REGION Network 19: QW98 - Spare Output (Hardware Channel De-activated)
   RUNG wire#powerrail
      P_Contact(operand := "80_From_HMI".MAN_AQ_INC_98, bit := "90_Manual_Data".INC_PLS_98)
      wire#w1
      Add(in1 := "16_AQ_Data".R2_SPR_AQ_98, in2 := 1.0, out => "16_AQ_Data".R2_SPR_AQ_98)
      { S7_Templates := "SrcType := Real" } GE_Contact(in1 := "16_AQ_Data".R2_SPR_AQ_98, in2 := "16_AQ_Data".QW_98.ENG_MAX)
      { S7_GenerateENO := "TRUE" } Move(in := "16_AQ_Data".QW_98.ENG_MAX, out1 => "16_AQ_Data".R2_SPR_AQ_98)
   END_RUNG
   RUNG wire#powerrail
      Contact( "80_From_HMI".MAN_AQ_INC_98 )
      P_Contact(operand := "Clock_5Hz", bit := "90_Manual_Data".INC_PLS_98_Hz)
   END_RUNG wire#w1
   RUNG wire#powerrail
      P_Contact(operand := "80_From_HMI".MAN_AQ_DEC_98, bit := "90_Manual_Data".DEC_PLS_98)
      wire#w2
      Sub(in1 := "16_AQ_Data".R2_SPR_AQ_98, in2 := 1.0, out => "16_AQ_Data".R2_SPR_AQ_98)
      { S7_Templates := "SrcType := Real" } LE_Contact(in1 := "16_AQ_Data".R2_SPR_AQ_98, in2 := "16_AQ_Data".QW_98.ENG_MIN)
      { S7_GenerateENO := "TRUE" } Move(in := "16_AQ_Data".QW_98.ENG_MIN, out1 => "16_AQ_Data".R2_SPR_AQ_98)
   END_RUNG
   RUNG wire#powerrail
      Contact( "80_From_HMI".MAN_AQ_DEC_98 )
      P_Contact(operand := "Clock_5Hz", bit := "90_Manual_Data".DEC_PLS_98_Hz)
   END_RUNG wire#w2
   // the same network as SCL:
   #_w1 := "80_From_HMI".MAN_AQ_INC_98 AND NOT "90_Manual_Data".INC_PLS_98;   // rising edge of "80_From_HMI".MAN_AQ_INC_98
   "90_Manual_Data".INC_PLS_98 := "80_From_HMI".MAN_AQ_INC_98;
   #_w2 := "80_From_HMI".MAN_AQ_INC_98 AND "Clock_5Hz" AND NOT "90_Manual_Data".INC_PLS_98_Hz;   // rising edge of "Clock_5Hz"
   "90_Manual_Data".INC_PLS_98_Hz := "Clock_5Hz";
   #_w3 := #_w1 OR #_w2;
   IF #_w3 THEN "16_AQ_Data".R2_SPR_AQ_98 := "16_AQ_Data".R2_SPR_AQ_98 + 1.0; END_IF;
   IF #_w3 AND ("16_AQ_Data".R2_SPR_AQ_98 >= "16_AQ_Data".QW_98.ENG_MAX) THEN
       "16_AQ_Data".R2_SPR_AQ_98 := "16_AQ_Data".QW_98.ENG_MAX;
   END_IF;
   #_w4 := "80_From_HMI".MAN_AQ_DEC_98 AND NOT "90_Manual_Data".DEC_PLS_98;   // rising edge of "80_From_HMI".MAN_AQ_DEC_98
   "90_Manual_Data".DEC_PLS_98 := "80_From_HMI".MAN_AQ_DEC_98;
   #_w5 := "80_From_HMI".MAN_AQ_DEC_98 AND "Clock_5Hz" AND NOT "90_Manual_Data".DEC_PLS_98_Hz;   // rising edge of "Clock_5Hz"
   "90_Manual_Data".DEC_PLS_98_Hz := "Clock_5Hz";
   #_w6 := #_w4 OR #_w5;
   IF #_w6 THEN "16_AQ_Data".R2_SPR_AQ_98 := "16_AQ_Data".R2_SPR_AQ_98 - 1.0; END_IF;
   IF #_w6 AND ("16_AQ_Data".R2_SPR_AQ_98 <= "16_AQ_Data".QW_98.ENG_MIN) THEN
       "16_AQ_Data".R2_SPR_AQ_98 := "16_AQ_Data".QW_98.ENG_MIN;
   END_IF;
END_REGION

REGION Network 20: QW100 - Main Fuel Reg Valve Control (CV-203)
   RUNG wire#powerrail
      P_Contact(operand := "80_From_HMI".MAN_AQ_INC_100, bit := "90_Manual_Data".INC_PLS_100)
      wire#w1
      Add(in1 := "16_AQ_Data".CV203_CNTRL, in2 := 1.0, out => "16_AQ_Data".CV203_CNTRL)
      { S7_Templates := "SrcType := Real" } GE_Contact(in1 := "16_AQ_Data".CV203_CNTRL, in2 := "16_AQ_Data".QW_100.ENG_MAX)
      { S7_GenerateENO := "TRUE" } Move(in := "16_AQ_Data".QW_100.ENG_MAX, out1 => "16_AQ_Data".CV203_CNTRL)
   END_RUNG
   RUNG wire#powerrail
      Contact( "80_From_HMI".MAN_AQ_INC_100 )
      P_Contact(operand := "Clock_5Hz", bit := "90_Manual_Data".INC_PLS_100_Hz)
   END_RUNG wire#w1
   RUNG wire#powerrail
      P_Contact(operand := "80_From_HMI".MAN_AQ_DEC_100, bit := "90_Manual_Data".DEC_PLS_100)
      wire#w2
      Sub(in1 := "16_AQ_Data".CV203_CNTRL, in2 := 1.0, out => "16_AQ_Data".CV203_CNTRL)
      { S7_Templates := "SrcType := Real" } LE_Contact(in1 := "16_AQ_Data".CV203_CNTRL, in2 := "16_AQ_Data".QW_100.ENG_MIN)
      { S7_GenerateENO := "TRUE" } Move(in := "16_AQ_Data".QW_100.ENG_MIN, out1 => "16_AQ_Data".CV203_CNTRL)
   END_RUNG
   RUNG wire#powerrail
      Contact( "80_From_HMI".MAN_AQ_DEC_100 )
      P_Contact(operand := "Clock_5Hz", bit := "90_Manual_Data".DEC_PLS_100_Hz)
   END_RUNG wire#w2
   // the same network as SCL:
   #_w1 := "80_From_HMI".MAN_AQ_INC_100 AND NOT "90_Manual_Data".INC_PLS_100;   // rising edge of "80_From_HMI".MAN_AQ_INC_100
   "90_Manual_Data".INC_PLS_100 := "80_From_HMI".MAN_AQ_INC_100;
   #_w2 := "80_From_HMI".MAN_AQ_INC_100 AND "Clock_5Hz" AND NOT "90_Manual_Data".INC_PLS_100_Hz;   // rising edge of "Clock_5Hz"
   "90_Manual_Data".INC_PLS_100_Hz := "Clock_5Hz";
   #_w3 := #_w1 OR #_w2;
   IF #_w3 THEN "16_AQ_Data".CV203_CNTRL := "16_AQ_Data".CV203_CNTRL + 1.0; END_IF;
   IF #_w3 AND ("16_AQ_Data".CV203_CNTRL >= "16_AQ_Data".QW_100.ENG_MAX) THEN
       "16_AQ_Data".CV203_CNTRL := "16_AQ_Data".QW_100.ENG_MAX;
   END_IF;
   #_w4 := "80_From_HMI".MAN_AQ_DEC_100 AND NOT "90_Manual_Data".DEC_PLS_100;   // rising edge of "80_From_HMI".MAN_AQ_DEC_100
   "90_Manual_Data".DEC_PLS_100 := "80_From_HMI".MAN_AQ_DEC_100;
   #_w5 := "80_From_HMI".MAN_AQ_DEC_100 AND "Clock_5Hz" AND NOT "90_Manual_Data".DEC_PLS_100_Hz;   // rising edge of "Clock_5Hz"
   "90_Manual_Data".DEC_PLS_100_Hz := "Clock_5Hz";
   #_w6 := #_w4 OR #_w5;
   IF #_w6 THEN "16_AQ_Data".CV203_CNTRL := "16_AQ_Data".CV203_CNTRL - 1.0; END_IF;
   IF #_w6 AND ("16_AQ_Data".CV203_CNTRL <= "16_AQ_Data".QW_100.ENG_MIN) THEN
       "16_AQ_Data".CV203_CNTRL := "16_AQ_Data".QW_100.ENG_MIN;
   END_IF;
END_REGION

REGION Network 21: QW102 - Main Atom Air Reg Valve Control (CV-111)
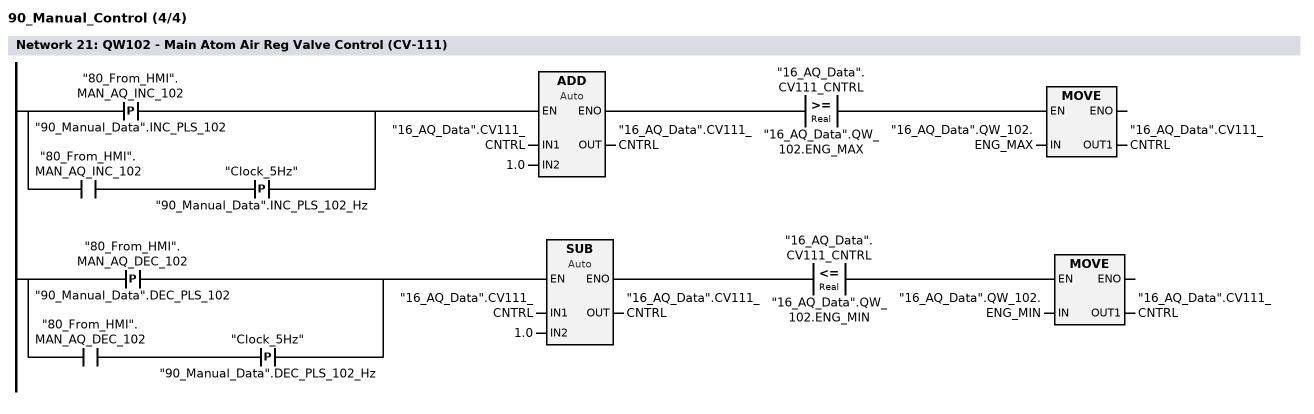
   RUNG wire#powerrail
      P_Contact(operand := "80_From_HMI".MAN_AQ_INC_102, bit := "90_Manual_Data".INC_PLS_102)
      wire#w1
      Add(in1 := "16_AQ_Data".CV111_CNTRL, in2 := 1.0, out => "16_AQ_Data".CV111_CNTRL)
      { S7_Templates := "SrcType := Real" } GE_Contact(in1 := "16_AQ_Data".CV111_CNTRL, in2 := "16_AQ_Data".QW_102.ENG_MAX)
      { S7_GenerateENO := "TRUE" } Move(in := "16_AQ_Data".QW_102.ENG_MAX, out1 => "16_AQ_Data".CV111_CNTRL)
   END_RUNG
   RUNG wire#powerrail
      Contact( "80_From_HMI".MAN_AQ_INC_102 )
      P_Contact(operand := "Clock_5Hz", bit := "90_Manual_Data".INC_PLS_102_Hz)
   END_RUNG wire#w1
   RUNG wire#powerrail
      P_Contact(operand := "80_From_HMI".MAN_AQ_DEC_102, bit := "90_Manual_Data".DEC_PLS_102)
      wire#w2
      Sub(in1 := "16_AQ_Data".CV111_CNTRL, in2 := 1.0, out => "16_AQ_Data".CV111_CNTRL)
      { S7_Templates := "SrcType := Real" } LE_Contact(in1 := "16_AQ_Data".CV111_CNTRL, in2 := "16_AQ_Data".QW_102.ENG_MIN)
      { S7_GenerateENO := "TRUE" } Move(in := "16_AQ_Data".QW_102.ENG_MIN, out1 => "16_AQ_Data".CV111_CNTRL)
   END_RUNG
   RUNG wire#powerrail
      Contact( "80_From_HMI".MAN_AQ_DEC_102 )
      P_Contact(operand := "Clock_5Hz", bit := "90_Manual_Data".DEC_PLS_102_Hz)
   END_RUNG wire#w2
   // the same network as SCL:
   #_w1 := "80_From_HMI".MAN_AQ_INC_102 AND NOT "90_Manual_Data".INC_PLS_102;   // rising edge of "80_From_HMI".MAN_AQ_INC_102
   "90_Manual_Data".INC_PLS_102 := "80_From_HMI".MAN_AQ_INC_102;
   #_w2 := "80_From_HMI".MAN_AQ_INC_102 AND "Clock_5Hz" AND NOT "90_Manual_Data".INC_PLS_102_Hz;   // rising edge of "Clock_5Hz"
   "90_Manual_Data".INC_PLS_102_Hz := "Clock_5Hz";
   #_w3 := #_w1 OR #_w2;
   IF #_w3 THEN "16_AQ_Data".CV111_CNTRL := "16_AQ_Data".CV111_CNTRL + 1.0; END_IF;
   IF #_w3 AND ("16_AQ_Data".CV111_CNTRL >= "16_AQ_Data".QW_102.ENG_MAX) THEN
       "16_AQ_Data".CV111_CNTRL := "16_AQ_Data".QW_102.ENG_MAX;
   END_IF;
   #_w4 := "80_From_HMI".MAN_AQ_DEC_102 AND NOT "90_Manual_Data".DEC_PLS_102;   // rising edge of "80_From_HMI".MAN_AQ_DEC_102
   "90_Manual_Data".DEC_PLS_102 := "80_From_HMI".MAN_AQ_DEC_102;
   #_w5 := "80_From_HMI".MAN_AQ_DEC_102 AND "Clock_5Hz" AND NOT "90_Manual_Data".DEC_PLS_102_Hz;   // rising edge of "Clock_5Hz"
   "90_Manual_Data".DEC_PLS_102_Hz := "Clock_5Hz";
   #_w6 := #_w4 OR #_w5;
   IF #_w6 THEN "16_AQ_Data".CV111_CNTRL := "16_AQ_Data".CV111_CNTRL - 1.0; END_IF;
   IF #_w6 AND ("16_AQ_Data".CV111_CNTRL <= "16_AQ_Data".QW_102.ENG_MIN) THEN
       "16_AQ_Data".CV111_CNTRL := "16_AQ_Data".QW_102.ENG_MIN;
   END_IF;
END_REGION
END_FUNCTION

// ===== PLC "Rack 3 - GCU & BWT PLC - 7KF2"  CPU 1516F-3 PN/DP =====

VAR_GLOBAL   // PLC tag table "Default tag table"
   "Clock_10Hz" AT %M0.0 : Bool;   // System bit
   "Clock_5Hz" AT %M0.1 : Bool;   // System bit
   "Clock_2.5Hz" AT %M0.2 : Bool;   // System bit
   "Clock_2Hz" AT %M0.3 : Bool;   // System bit
   "Clock_1.25Hz" AT %M0.4 : Bool;   // System bit
   "Clock_1Hz" AT %M0.5 : Bool;   // System bit
   "Clock_0.625Hz" AT %M0.6 : Bool;   // System bit
   "Clock_0.5Hz" AT %M0.7 : Bool;   // System bit
   "Clock_Byte" AT %MB0 : Byte;   // System bit
   "System_Byte" AT %MB1 : Byte;   // System bit
   "FirstScan" AT %M1.0 : Bool;   // System bit
   "DiagStatusUpdate" AT %M1.1 : Bool;   // System bit
   "AlwaysTRUE" AT %M1.2 : Bool;   // System bit
   "AlwaysFALSE" AT %M1.3 : Bool;   // System bit
   "Tag_1" AT %M222.2 : Bool;
   "Tag_2" AT %ID222 : Real;
   "Tag_3" AT %ID223 : Real;
   "Tag_4" AT %ID224 : Real;
   "Tag_5" AT %ID221 : Real;
   "Tag_6" AT %M1000.0 : Bool;
   "Tag_7" AT %MD1002 : Real;
   "TEST" AT %M2.0 : Bool;
   "Tag_8" AT %M55.0 : Bool;
   "Tag_9" AT %MD55 : DWord;
   "Tag_10" AT %MD56 : Real;
   "Tag_11" AT %MD57 : Real;
   "Tag_12" AT %MD58 : DWord;
   "Tag_13" AT %MD59 : Real;
   "Tag_14" AT %MD60 : DWord;
   "Tag_15" AT %MD61 : Real;
   "Tag_16" AT %MD62 : DWord;
   "Tag_17" AT %MD63 : Real;
   "Tag_18" AT %MD64 : DWord;
   "Tag_19" AT %MD65 : Real;
   "Tag_20" AT %MD66 : DWord;
   "Tag_21" AT %MD67 : Real;
   "Tag_22" AT %MD68 : DWord;
   "Tag_23" AT %MD69 : DWord;
   "Tag_24" AT %MD70 : Real;
   "Tag_25" AT %MD71 : DWord;
   "Tag_26" AT %MD72 : Real;
   "Tag_27" AT %MD73 : Real;
   "Tag_28" AT %MD74 : DWord;
   "Tag_29" AT %MD75 : Real;
   "Tag_30" AT %MD76 : DWord;
   "Tag_31" AT %MD77 : Real;
   "Tag_32" AT %MD78 : DWord;
   "Tag_33" AT %MD79 : Real;
   "Tag_34" AT %MD80 : DWord;
   "Tag_35" AT %MD81 : Real;
   "Tag_36" AT %MD82 : DWord;
END_VAR

VAR_GLOBAL   // PLC tag table "PLC_IO"
   "R3_SPR_DI_136_0" AT %I136.0 : Bool;   // Spare input
   "R3_SPR_DI_136_1" AT %I136.1 : Bool;   // Spare input
   "Cooling Seawater Flow Switch" AT %I136.2 : Bool;   // FS332-8B1
   "Fresh Water Cooling Flow Switch" AT %I136.5 : Bool;   // FS350-8B3
   "GCU Drain Valve Feedback Open" AT %I136.6 : Bool;   // CV341-8B4
   "GCU Drain Valve Feedback Closed" AT %I136.7 : Bool;   // CV341-8B4
   "Gas to Deck Valve Feedback Open" AT %I137.0 : Bool;   // CV406-9B1
   "Gas to Deck Valve Feedback Closed" AT %I137.1 : Bool;   // CV406-9B1
   "Gas Block Valve 1 Feedback Open" AT %I137.2 : Bool;   // CV407-9B2
   "Gas Block Valve 1 Feedback Closed" AT %I137.3 : Bool;   // CV407-9B2
   "Gas Block Valve 2 Feedback Open" AT %I137.4 : Bool;   // CV411-9B3
   "Gas Block Valve 2 Feedback Closed" AT %I137.5 : Bool;   // CV411-9B3
   "Gas Bleed Valve Feedback Open" AT %I137.6 : Bool;   // CV409-9B4
   "Gas Bleed Valve Feedback Closed" AT %I137.7 : Bool;   // CV409-9B4
   "Ambient Air Valve Feedback Open" AT %I138.0 : Bool;   // CV441-10B1
   "Ambient Air Valve Feedback Closed" AT %I138.1 : Bool;   // CV441-10B1
   "GCU Low Level Switch" AT %I138.2 : Bool;   // LS303-10B2
   "GCU Booster Pump Enabled" AT %I138.3 : Bool;   // P304-MCCP
   "GCU Local PB - Start" AT %I138.4 : Bool;   // 10S1
   "GCU Local PB - Stop" AT %I138.5 : Bool;   // 10S2
   "E-Stop Pressed @ BWT CP" AT %I138.6 : Bool;   // 8S1
   "GCU Recirculation Pump Enabled" AT %I138.7 : Bool;   // P303-MCCP
   "Process Gas Compressor Running/Stopped" AT %I139.0 : Bool;   // E400
   "Process Gas Compressor Tripped/Shutdown" AT %I139.1 : Bool;   // E400
   "GCU Recirculation Pump Healthy" AT %I139.2 : Bool;   // P303-MCCP
   "5T1 Power Healthy" AT %I139.3 : Bool;   // 5T2
   "Panel Vent Power Healthy" AT %I139.4 : Bool;   // 6Q6
   "GCU Booster Pump Healthy" AT %I139.5 : Bool;   // P304-MCCP
   "PGC Running Loaded/On-line" AT %I139.6 : Bool;   // E400
   "PGC Alarm/Warning" AT %I139.7 : Bool;   // E400
   "GCU Level" AT %IW800 : Int;   // LIT304
   "R3_SPR_AI_802" AT %IW802 : Int;   // Spare input
   "Fresh Water Cooling Temperature" AT %IW804 : Int;   // TIT408
   "Gas to Deck (Outlet) Temperature" AT %IW806 : Int;   // TIT406
   "Gas To Deck Vent Valve Feedback" AT %IW808 : Int;   // CV405
   "Gas to Deck Pressure" AT %IW810 : Int;   // PIT416
   "Fresh Water Inlet Pressure" AT %IW812 : Int;   // PIT358
   "GCU Cooling Seawater Pressure" AT %IW814 : Int;   // PIT348
   "Recirculation Fresh Water Pressure" AT %IW816 : Int;   // PIT353
   "PGC Discharge (outlet) Pressure" AT %IW818 : Int;   // E400-PT002
   "PGC Discharge (Outlet) Temperature" AT %IW820 : Int;   // E400-TT002
   "Ballast Water Salinity" AT %IW822 : Int;   // SL-400
   "R3_SPR_AI_824" AT %IW824 : Int;   // Spare input
   "R3_SPR_AI_826" AT %IW826 : Int;   // Spare input
   "R3_SPR_AI_828" AT %IW828 : Int;   // Spare input
   "R3_SPR_AI_830" AT %IW830 : Int;   // Spare input
   "Fresh Water Fill Valve Control" AT %Q136.0 : Bool;   // CV358 / 12QM1
   "Waste Water Drain Valve Control" AT %Q136.1 : Bool;   // CV341 / 12QM2
   "Block Valve 1 Control" AT %Q136.2 : Bool;   // CV407 / 12QM3
   "Bleed Valve Control" AT %Q136.3 : Bool;   // CV409 / 12QM4
   "Block Valve 2 Control" AT %Q136.4 : Bool;   // CV411 / 12QM5
   "Ambient Air Valve Control" AT %Q136.5 : Bool;   // CV441 / 12QM6
   "Main Gas to Deck Valve Control" AT %Q136.6 : Bool;   // CV406 / 12QM7
   "Start Process Gas Compressor" AT %Q136.7 : Bool;   // E400-Start
   "GCU Recirculation Pump Control" AT %Q137.0 : Bool;   // P303
   "GCU Booster Pump Control" AT %Q137.1 : Bool;   // P304
   "GCU Warning Alarm" AT %Q137.2 : Bool;   // 13P1
   "GCU Shutdown Alarm" AT %Q137.3 : Bool;   // 13P2
   "GCU Running" AT %Q137.4 : Bool;   // 13P3
   "Ballast Water Tank Level High High" AT %Q137.5 : Bool;   // 13P4
   "GCU Alarm Buzzer" AT %Q137.6 : Bool;   // 13P5
   "Stop Process Gas Compressor" AT %Q137.7 : Bool;   // E400-Stop
   "Pilot For GTT FPT Valve" AT %Q138.0 : Bool;   // CV422-FPT / 14QM1
   "Pilot For GTT 1 Port Valve" AT %Q138.1 : Bool;   // CV422-1P / 14QM2
   "Pilot For GTT 1 Starboard Valve" AT %Q138.2 : Bool;   // CV421-1S / 14QM3
   "Pilot For GTT 2 Port Valve" AT %Q138.3 : Bool;   // CV422-2P / 14QM4
   "Pilot For GTT 2 Starboard Valve" AT %Q138.4 : Bool;   // CV421-2S / 14QM5
   "Pilot For GTT 3 Port Valve" AT %Q138.5 : Bool;   // CV422-3P / 14QM6
   "Pilot For GTT 3 Starboard Valve" AT %Q138.6 : Bool;   // CV421-3S / 14QM7
   "R3_SPR_DQ_138_7" AT %Q138.7 : Bool;   // Spare output
   "Pilot For GTT 4 Port Valve" AT %Q139.0 : Bool;   // CV422-4P / 15QM1
   "Pilot For GTT 4 Starboard Valve" AT %Q139.1 : Bool;   // CV421-4S / 15QM2
   "Pilot For GTT 5 Port Valve" AT %Q139.2 : Bool;   // CV422-5P / 15QM3
   "Pilot For GTT 5 Starboard Valve" AT %Q139.3 : Bool;   // CV421-5S / 15QM4
   "Pilot For GTT 6 Port Valve" AT %Q139.4 : Bool;   // CV422-6P / 15QM5
   "Pilot For GTT 6 Starboard Valve" AT %Q139.5 : Bool;   // CV421-6S / 15QM6
   "Pilot For GTT APT Port Valve" AT %Q139.6 : Bool;   // CV422-APT / 15QM7
   "R3_SPR_DQ_139_7" AT %Q139.7 : Bool;   // Spare output
   "Gas Vent Position Control" AT %QW800 : Int;   // CV405
   "R3_SPR_AQ_802" AT %QW802 : Int;   // Spare output
   "R3_SPR_AQ_804" AT %QW804 : Int;   // Spare output
   "R3_SPR_AQ_806" AT %QW806 : Int;   // Spare output
   "FW Fill Valve Feedback Closed" AT %I136.4 : Bool;   // CV358-8B2
   "FW Fill Valve Feedback Open" AT %I136.3 : Bool;   // CV358-8B2
END_VAR

VAR_GLOBAL   // PLC tag table "RIO_1"
   "FPT USD Flow Meter" AT %IW100 : Int;   // FIT418-FPT
   "FPT MBG Flow Meter" AT %IW102 : Int;   // FIT420-FPT
   "Tank 1P USD Flow Meter" AT %IW104 : Int;   // FIT418-1P
   "Tank 1P MBG Flow Meter" AT %IW106 : Int;   // FIT420-1P
   "Tank 1S USD Flow Meter" AT %IW108 : Int;   // FIT417-1S
   "Tank 1S MBG Flow Meter" AT %IW110 : Int;   // FIT419-1S
   "RIO1_SPR_AI_114" AT %IW114 : Int;   // Spare input
   "FPT BWT Level" AT %IW118 : Int;   // LT422-FPT
   "Tank 1P BWT Level" AT %IW120 : Int;   // LT422-1P
   "Tank 1S BWT Level" AT %IW122 : Int;   // LT421-1S
   "FPT BWT ph" AT %IW124 : Int;   // 426-FPT
   "FPT BWT Temp" AT %IW126 : Int;   // 426-FPT
   "FPT BWT DO" AT %IW128 : Int;   // 428-FPT
   "Tank 1S BWT ph" AT %IW140 : Int;   // 425-1S
   "Tank 1S BWT Temp" AT %IW142 : Int;   // 425-1S
   "Tank 1S BWT DO" AT %IW144 : Int;   // 427-1S
   "RIO1_SPR_AI_146" AT %IW146 : Int;   // Spare input
   "Tank 1P BWT ph" AT %IW148 : Int;   // 426-1P
   "Tank 1P BWT Temp" AT %IW150 : Int;   // 426-1P
   "Tank 1P BWT DO" AT %IW152 : Int;   // 428-1P
   "RIO1_SPR_AI_154" AT %IW154 : Int;   // Spare input
   "FPT GTT Isolation Valve Feedback - Opened" AT %I0.0 : Bool;   // CV422
   "FPT GTT Isolation Valve Feedback - Closed" AT %I0.1 : Bool;   // CV422
   "FPT Tank Vent Valve 1 Feedback - Opened" AT %I0.2 : Bool;   // CV441-FPTA
   "FPT Tank Vent Valve 1 Feedback - Closed" AT %I0.3 : Bool;   // CV441-FPTA
   "FPT Tank Vent Valve 2 Feedback - Opened" AT %I0.4 : Bool;   // CV441-FPTB
   "FPT Tank Vent Valve 2 Feedback - Closed" AT %I0.5 : Bool;   // CV441-FPTB
   "RIO1_SPR_DI_0_6" AT %I0.6 : Bool;   // Spare input
   "RIO1_SPR_DI_0_7" AT %I0.7 : Bool;   // Spare input
   "Tank 1P GTT Isolation Valve Feedback - Opened" AT %I3.0 : Bool;   // CV422
   "Tank 1P GTT Isolation Valve Feedback - Closed" AT %I3.1 : Bool;   // CV422
   "Tank 1P Tank Vent Valve 1 Feedback - Opened" AT %I3.2 : Bool;   // CV441-1PA
   "Tank 1P Tank Vent Valve 1 Feedback - Closed" AT %I3.3 : Bool;   // CV441-1PA
   "Tank 1P Tank Vent Valve 2 Feedback - Opened" AT %I3.4 : Bool;   // CV441-1PB
   "Tank 1P Tank Vent Valve 2 Feedback - Closed" AT %I3.5 : Bool;   // CV441-1PB
   "RIO1_SPR_DI_3_6" AT %I3.6 : Bool;   // Spare input
   "RIO1_SPR_DI_3_7" AT %I3.7 : Bool;   // Spare input
   "Tank 1S GTT Isolation Valve Feedback - Opened" AT %I6.0 : Bool;   // CV421
   "Tank 1S GTT Isolation Valve Feedback - Closed" AT %I6.1 : Bool;   // CV421
   "Tank 1S Tank Vent Valve 1 Feedback - Opened" AT %I6.2 : Bool;   // CV440-1SA
   "Tank 1S Tank Vent Valve 1 Feedback - Closed" AT %I6.3 : Bool;   // CV440-1SA
   "Tank 1S Tank Vent Valve 2 Feedback - Opened" AT %I6.4 : Bool;   // CV440-1SB
   "Tank 1S Tank Vent Valve 2 Feedback - Closed" AT %I6.5 : Bool;   // CV440-1SB
   "RIO1_SPR_DI_6_6" AT %I6.6 : Bool;   // Spare input
   "RIO1_SPR_DI_6_7" AT %I6.7 : Bool;   // Spare input
   "FPT BWT Level High High Switch" AT %I9.0 : Bool;   // LS425-FPT
   "RIO1 Tanks Pressure Switch Hi Hi" AT %I9.1 : Bool;   // PS436-FPT/1P/1S
   "Tank 1P BWT Level High High Switch" AT %I9.2 : Bool;   // LS425-1P
   "Tank 1S BWT Level High High Switch" AT %I9.3 : Bool;   // LS425-1S
   "RIO1_SPR_DI_9_4" AT %I9.4 : Bool;   // Spare input
   "RIO1_SPR_DI_9_5" AT %I9.5 : Bool;   // Spare input
   "RIO1_SPR_DI_9_6" AT %I9.6 : Bool;   // Spare input
   "RIO1_SPR_DI_9_7" AT %I9.7 : Bool;   // Spare input
   "FTP Vent Valve 1" AT %Q0.0 : Bool;   // CV441-FPTA
   "FTP Vent Valve 2" AT %Q0.1 : Bool;   // CV441-FPTB
   "Tank 1P Vent Valve 1" AT %Q0.2 : Bool;   // CV441-1PA
   "Tank 1P Vent Valve 2" AT %Q0.3 : Bool;   // CV441-1PB
   "Tank 1S Vent Valve 1" AT %Q2.0 : Bool;   // CV440-1SA
   "Tank 1S Vent Valve 2" AT %Q2.1 : Bool;   // CV440-1SB
   "RIO1 Confined Space O2 Monitor" AT %IW112 : Int;   // 600-TX-433
   "RIO1 Deck Main IG Pressure Transmitter" AT %IW116 : Int;   // PT415
   "RIO1 Tanks Pressure Transmitter" AT %IW130 : Int;   // PT424-FPT/1P/1S
   "RIO1_SPR_DQ_2_2" AT %Q2.2 : Bool;   // Spare output
   "RIO1_SPR_DQ_2_3" AT %Q2.3 : Bool;   // Spare output
END_VAR

VAR_GLOBAL   // PLC tag table "RIO_2"
   "Tank 2P GTT Isolation Valve Feedback - Opened" AT %I15.0 : Bool;   // CV422-2P
   "Tank 2P GTT Isolation Valve Feedback - Closed" AT %I15.1 : Bool;   // CV422-2P
   "Tank 2P Tank Vent Valve 1 Feedback - Opened" AT %I15.2 : Bool;   // CV441-2P1
   "Tank 2P Tank Vent Valve 1 Feedback - Closed" AT %I15.3 : Bool;   // CV441-2P1
   "Tank 2P Tank Vent Valve 2 Feedback - Opened" AT %I15.4 : Bool;   // CV441-2P2
   "Tank 2P Tank Vent Valve 2 Feedback - Closed" AT %I15.5 : Bool;   // CV441-2P2
   "RIO2_SPR_DI_15_6" AT %I15.6 : Bool;   // Spare input
   "RIO2_SPR_DI_15_7" AT %I15.7 : Bool;   // Spare input
   "Tank 2S GTT Isolation Valve Feedback - Opened" AT %I18.0 : Bool;   // CV421-2S
   "Tank 2S GTT Isolation Valve Feedback - Closed" AT %I18.1 : Bool;   // CV421-2S
   "Tank 2S Tank Vent Valve 1 Feedback - Opened" AT %I18.2 : Bool;   // CV440-2SA
   "Tank 2S Tank Vent Valve 1 Feedback - Closed" AT %I18.3 : Bool;   // CV440-2SA
   "Tank 2S Tank Vent Valve 2 Feedback - Opened" AT %I18.4 : Bool;   // CV440-2SB
   "Tank 2S Tank Vent Valve 2 Feedback - Closed" AT %I18.5 : Bool;   // CV440-2SB
   "RIO2_SPR_DI_18_6" AT %I18.6 : Bool;   // Spare input
   "RIO2_SPR_DI_18_7" AT %I18.7 : Bool;   // Spare input
   "Tank 2P BWT Level High High Switch" AT %I21.0 : Bool;   // LS425-2P
   "RIO2 Tanks Pressure Switch Hi Hi" AT %I21.1 : Bool;   // PS436-2P/2S
   "Tank 2S BWT Level High High Switch" AT %I21.2 : Bool;   // LS422-2S
   "RIO2_SPR_DI_21_3" AT %I21.3 : Bool;   // Spare input
   "RIO2_SPR_DI_21_4" AT %I21.4 : Bool;   // Spare input
   "RIO2_SPR_DI_21_5" AT %I21.5 : Bool;   // Spare input
   "RIO2_SPR_DI_21_6" AT %I21.6 : Bool;   // Spare input
   "RIO2_SPR_DI_21_7" AT %I21.7 : Bool;   // Spare input
   "Tank 2P USD Flow Meter" AT %IW160 : Int;   // FIT418-2P
   "Tank 2P MBG Flow Meter" AT %IW162 : Int;   // FIT420-2P
   "Tank 2S USD Flow Meter" AT %IW164 : Int;   // FIT417-2S
   "Tank 2S MBG Flow Meter" AT %IW166 : Int;   // FIT419-2S
   "RIO2 Main Gas-To-Deck Pressure" AT %IW168 : Int;   // PT415
   "Tank 2P BWT Level" AT %IW170 : Int;   // LT422-2P
   "Tank 2S BWT Level" AT %IW172 : Int;   // LT421-2S
   "RIO2_SPR_AI_174" AT %IW174 : Int;   // Spare input
   "Tank 2P BWT ph" AT %IW176 : Int;   // 426-2P
   "Tank 2P BWT Temp" AT %IW178 : Int;   // 426-2P
   "Tank 2P BWT DO" AT %IW180 : Int;   // 428-2P
   "RIO2 Tanks Pressure" AT %IW182 : Int;   // PT424-2P/2S
   "Tank 2S BWT ph" AT %IW184 : Int;   // 425-2S
   "Tank 2S BWT Temp" AT %IW186 : Int;   // 425-2S
   "Tank 2S BWT DO" AT %IW188 : Int;   // 427-2S
   "RIO2 Confined Space O2 Monitor" AT %IW190 : Int;   // 600-TX-433
   "Tank 2P Vent Valve 1" AT %Q6.0 : Bool;   // CV441-2PA
   "Tank 2P Vent Valve 2" AT %Q6.1 : Bool;   // CV441-2PA
   "Tank 2S Vent Valve 1" AT %Q6.2 : Bool;   // CV440-2SA
   "Tank 2S Vent Valve 2" AT %Q6.3 : Bool;   // CV440-2SA
END_VAR

VAR_GLOBAL   // PLC tag table "RIO_3"
   "Tank 3P GTT Isolation Valve Feedback - Opened" AT %I27.0 : Bool;   // CV422-3P
   "Tank 3P GTT Isolation Valve Feedback - Closed" AT %I27.1 : Bool;   // CV422-3P
   "Tank 3P Tank Vent Valve 1 Feedback - Opened" AT %I27.2 : Bool;   // CV441-3PA
   "Tank 3P Tank Vent Valve 1 Feedback - Closed" AT %I27.3 : Bool;   // CV441-3PA
   "Tank 3P Tank Vent Valve 2 Feedback - Opened" AT %I27.4 : Bool;   // CV441-3PB
   "Tank 3P Tank Vent Valve 2 Feedback - Closed" AT %I27.5 : Bool;   // CV441-3PB
   "RIO3_SPR_DI_27_6" AT %I27.6 : Bool;   // Spare input
   "RIO3_SPR_DI_27_7" AT %I27.7 : Bool;   // Spare input
   "Tank 3S GTT Isolation Valve Feedback - Opened" AT %I30.0 : Bool;   // CV421-3S
   "Tank 3S GTT Isolation Valve Feedback - Closed" AT %I30.1 : Bool;   // CV421-3S
   "Tank 3S Tank Vent Valve 1 Feedback - Opened" AT %I30.2 : Bool;   // CV440-3SA
   "Tank 3S Tank Vent Valve 1 Feedback - Closed" AT %I30.3 : Bool;   // CV440-3SA
   "Tank 3S Tank Vent Valve 2 Feedback - Opened" AT %I30.4 : Bool;   // CV440-3SB
   "Tank 3S Tank Vent Valve 2 Feedback - Closed" AT %I30.5 : Bool;   // CV440-3SB
   "RIO3_SPR_DI_30_6" AT %I30.6 : Bool;   // Spare input
   "RIO3_SPR_DI_30_7" AT %I30.7 : Bool;   // Spare input
   "Tank 3P BWT Level High High Switch" AT %I33.0 : Bool;   // LS425-3P
   "RIO3 Tanks Pressure Switch Hi Hi" AT %I33.1 : Bool;   // PS436-3P/3S
   "Tank 3S BWT Level High High Switch" AT %I33.2 : Bool;   // LS422-3S
   "RIO3_SPR_DI_33_3" AT %I33.3 : Bool;   // Spare input
   "RIO3_SPR_DI_33_4" AT %I33.4 : Bool;   // Spare input
   "RIO3_SPR_DI_33_5" AT %I33.5 : Bool;   // Spare input
   "RIO3_SPR_DI_33_6" AT %I33.6 : Bool;   // Spare input
   "RIO3_SPR_DI_33_7" AT %I33.7 : Bool;   // Spare input
   "Tank 3P USD Flow Meter" AT %IW200 : Int;   // FIT418-3P
   "Tank 3P MBG Flow Meter" AT %IW202 : Int;   // FIT420-3P
   "Tank 3S USD Flow Meter" AT %IW204 : Int;   // FIT417-3S
   "Tank 3S MBG Flow Meter" AT %IW206 : Int;   // FIT419-3S
   "RIO3 Main Gas-To-Deck Pressure" AT %IW208 : Int;   // PT415
   "Tank 3P BWT Level" AT %IW210 : Int;   // LT422-3P
   "Tank 3S BWT Level" AT %IW212 : Int;   // LT421-3S
   "RIO3_SPR_AI_214" AT %IW214 : Int;   // Spare input
   "Tank 3P BWT ph" AT %IW216 : Int;   // 426-3P
   "Tank 3P BWT Temp" AT %IW218 : Int;   // 426-3P
   "Tank 3P BWT DO" AT %IW220 : Int;   // 428-3P
   "RIO3 Tanks Pressure" AT %IW222 : Int;   // PT424-3P/3S
   "Tank 3S BWT ph" AT %IW224 : Int;   // 425-3S
   "Tank 3S BWT Temp" AT %IW226 : Int;   // 425-3S
   "Tank 3S BWT DO" AT %IW228 : Int;   // 427-3S
   "RIO3_SPR_AI_230" AT %IW230 : Int;   // Spare input
   "Tank 3P Vent Valve 1" AT %Q10.0 : Bool;   // CV441-3PA
   "Tank 3P Vent Valve 2" AT %Q10.1 : Bool;   // CV441-3PB
   "Tank 3S Vent Valve 1" AT %Q10.2 : Bool;   // CV440-3SA
   "Tank 3S Vent Valve 2" AT %Q10.3 : Bool;   // CV440-3SB
END_VAR

VAR_GLOBAL   // PLC tag table "RIO_4"
   "Tank 4P GTT Isolation Valve Feedback - Opened" AT %I39.0 : Bool;   // CV422-4P
   "Tank 4P GTT Isolation Valve Feedback - Closed" AT %I39.1 : Bool;   // CV422-4P
   "Tank 4P Tank Vent Valve 1 Feedback - Opened" AT %I39.2 : Bool;   // CV441-4PA
   "Tank 4P Tank Vent Valve 1 Feedback - Closed" AT %I39.3 : Bool;   // CV441-4PA
   "Tank 4P Tank Vent Valve 2 Feedback - Opened" AT %I39.4 : Bool;   // CV441-4PB
   "Tank 4P Tank Vent Valve 2 Feedback - Closed" AT %I39.5 : Bool;   // CV441-4PB
   "RIO4_SPR_DI_139_6" AT %I39.6 : Bool;   // Spare input
   "RIO4_SPR_DI_139_7" AT %I39.7 : Bool;   // Spare input
   "Tank 4S GTT Isolation Valve Feedback - Opened" AT %I42.0 : Bool;   // CV421-4S
   "Tank 4S GTT Isolation Valve Feedback - Closed" AT %I42.1 : Bool;   // CV421-4S
   "Tank 4S Tank Vent Valve 1 Feedback - Opened" AT %I42.2 : Bool;   // CV440-4SA
   "Tank 4S Tank Vent Valve 1 Feedback - Closed" AT %I42.3 : Bool;   // CV440-4SA
   "Tank 4S Tank Vent Valve 2 Feedback - Opened" AT %I42.4 : Bool;   // CV440-4SB
   "Tank 4S Tank Vent Valve 2 Feedback - Closed" AT %I42.5 : Bool;   // CV440-4SB
   "RIO4_SPR_DI_142_6" AT %I42.6 : Bool;   // Spare input
   "RIO4_SPR_DI_142_7" AT %I42.7 : Bool;   // Spare input
   "Tank 4P BWT Level High High Switch" AT %I45.0 : Bool;   // LS425-4P
   "RIO4 Tanks Pressure Switch Hi Hi" AT %I45.1 : Bool;   // PS436-4P/4S
   "Tank 4S BWT Level High High Switch" AT %I45.2 : Bool;   // LS422-4S
   "RIO4_SPR_DI_145_3" AT %I45.3 : Bool;   // Spare input
   "RIO4_SPR_DI_145_4" AT %I45.4 : Bool;   // Spare input
   "RIO4_SPR_DI_145_5" AT %I45.5 : Bool;   // Spare input
   "RIO4_SPR_DI_145_6" AT %I45.6 : Bool;   // Spare input
   "RIO4_SPR_DI_145_7" AT %I45.7 : Bool;   // Spare input
   "Tank 4P USD Flow Meter" AT %IW260 : Int;   // FIT418-4P
   "Tank 4P MBG Flow Meter" AT %IW262 : Int;   // FIT420-4P
   "Tank 4S USD Flow Meter" AT %IW264 : Int;   // FIT417-4S
   "Tank 4S MBG Flow Meter" AT %IW266 : Int;   // FIT419-4S
   "RIO4 Main Gas-To-Deck Pressure" AT %IW268 : Int;   // PT415
   "Tank 4P BWT Level" AT %IW270 : Int;   // LT422-4P
   "Tank 4S BWT Level" AT %IW272 : Int;   // LT421-4S
   "RIO4_SPR_AI_274" AT %IW274 : Int;   // Spare input
   "Tank 4P BWT ph" AT %IW276 : Int;   // 426-4P
   "Tank 4P BWT Temp" AT %IW278 : Int;   // 426-4P
   "Tank 4P BWT DO" AT %IW280 : Int;   // 428-4P
   "RIO4 Tanks Pressure" AT %IW282 : Int;   // PT424-4P/4S
   "Tank 4S BWT ph" AT %IW284 : Int;   // 425-4S
   "Tank 4S BWT Temp" AT %IW286 : Int;   // 425-4S
   "Tank 4S BWT DO" AT %IW288 : Int;   // 427-4S
   "RIO4_SPR_AI_290" AT %IW290 : Int;   // Spare input
   "Tank 4P Vent Valve 1" AT %Q14.0 : Bool;   // CV441-4PA
   "Tank 4P Vent Valve 2" AT %Q14.1 : Bool;   // CV441-4PB
   "Tank 4S Vent Valve 1" AT %Q14.2 : Bool;   // CV440-4SA
   "Tank 4S Vent Valve 2" AT %Q14.3 : Bool;   // CV440-4SB
END_VAR

VAR_GLOBAL   // PLC tag table "RIO_5"
   "Tank 5P GTT Isolation Valve Feedback - Opened" AT %I51.0 : Bool;   // CV422-5P
   "Tank 5P GTT Isolation Valve Feedback - Closed" AT %I51.1 : Bool;   // CV422-5P
   "Tank 5P Tank Vent Valve 1 Feedback - Opened" AT %I51.2 : Bool;   // CV441-5PA
   "Tank 5P Tank Vent Valve 1 Feedback - Closed" AT %I51.3 : Bool;   // CV441-5PA
   "Tank 5P Tank Vent Valve 2 Feedback - Opened" AT %I51.4 : Bool;   // CV441-5PB
   "Tank 5P Tank Vent Valve 2 Feedback - Closed" AT %I51.5 : Bool;   // CV441-5PB
   "RIO5_SPR_DI_51_6" AT %I51.6 : Bool;   // Spare input
   "RIO5_SPR_DI_51_7" AT %I51.7 : Bool;   // Spare input
   "Tank 5S GTT Isolation Valve Feedback - Opened" AT %I54.0 : Bool;   // CV421-5S
   "Tank 5S GTT Isolation Valve Feedback - Closed" AT %I54.1 : Bool;   // CV421-5S
   "Tank 5S Tank Vent Valve 1 Feedback - Opened" AT %I54.2 : Bool;   // CV440-5SA
   "Tank 5S Tank Vent Valve 1 Feedback - Closed" AT %I54.3 : Bool;   // CV440-5SA
   "Tank 5S Tank Vent Valve 2 Feedback - Opened" AT %I54.4 : Bool;   // CV440-5SB
   "Tank 5S Tank Vent Valve 2 Feedback - Closed" AT %I54.5 : Bool;   // CV440-5SB
   "RIO5_SPR_DI_54_6" AT %I54.6 : Bool;   // Spare input
   "RIO5_SPR_DI_54_7" AT %I54.7 : Bool;   // Spare input
   "Tank 5P BWT Level High High Switch" AT %I57.0 : Bool;   // LS425-5P
   "RIO5 Tanks Pressure Switch Hi Hi" AT %I57.1 : Bool;   // PS436-5P/5S
   "Tank 5S BWT Level High High Switch" AT %I57.2 : Bool;   // LS422-5S
   "RIO5_SPR_DI_57_3" AT %I57.3 : Bool;   // Spare input
   "RIO5_SPR_DI_57_4" AT %I57.4 : Bool;   // Spare input
   "RIO5_SPR_DI_57_5" AT %I57.5 : Bool;   // Spare input
   "RIO5_SPR_DI_57_6" AT %I57.6 : Bool;   // Spare input
   "RIO5_SPR_DI_57_7" AT %I57.7 : Bool;   // Spare input
   "Tank 5P USD Flow Meter" AT %IW300 : Int;   // FIT418-5P
   "Tank 5P MBG Flow Meter" AT %IW302 : Int;   // FIT420-5P
   "Tank 5S USD Flow Meter" AT %IW304 : Int;   // FIT417-5S
   "Tank 5S MBG Flow Meter" AT %IW306 : Int;   // FIT419-5S
   "RIO5 Main Gas-To-Deck Pressure" AT %IW308 : Int;   // PT415
   "Tank 5P BWT Level" AT %IW310 : Int;   // LT422-5P
   "Tank 5S BWT Level" AT %IW312 : Int;   // LT421-5S
   "RIO5_SPR_AI_314" AT %IW314 : Int;   // Spare input
   "Tank 5P BWT ph" AT %IW316 : Int;   // 426-5P
   "Tank 5P BWT Temp" AT %IW318 : Int;   // 426-5P
   "Tank 5P BWT DO" AT %IW320 : Int;   // 428-5P
   "RIO5 Tanks Pressure" AT %IW322 : Int;   // PT424-5P/5S
   "Tank 5S BWT ph" AT %IW324 : Int;   // 425-5S
   "Tank 5S BWT Temp" AT %IW326 : Int;   // 425-5S
   "Tank 5S BWT DO" AT %IW328 : Int;   // 427-5S
   "RIO5_SPR_AI_330" AT %IW330 : Int;   // Spare input
   "Tank 5P Vent Valve 1" AT %Q18.0 : Bool;   // CV441-5PA
   "Tank 5P Vent Valve 2" AT %Q18.1 : Bool;   // CV441-5PA
   "Tank 5S Vent Valve 1" AT %Q18.2 : Bool;   // CV440-5SA
   "Tank 5S Vent Valve 2" AT %Q18.3 : Bool;   // CV440-5SA
END_VAR
